
       ELSE

           "Z256_Manager".tOutputData.dMissionCode := "Z256_Manager".tInputData.dMissionCode;
           "Z256_Manager".tOutputData.rgxFireHeadON_OFF := "Z256_Manager".tInputData.rgxFireRequest;
           FOR #TMP_dIndex2 := 0 TO "CONST_dNumberOfHeadsCycle" DO
               "Z256_Manager".tOutputData.rgxDataToProcessInter[#TMP_dIndex2] := true;
           END_FOR;
           "Z256_Manager".tOutputData.dTargetLineValue_cmm := "Z256_Manager".tInputData.dMissionStart_cmm;

           #TMP_iReturn := "GP_BlockMoveStruct"(IN_iCount := DINT_TO_INT("CONST_dNumberOfHeads"),
                                                IN_iDestIndex := 0,
                                                IN_iSourceIndex := 0,
                                                INO_vDestArrayStruct := "Z256_Manager".tOutputData.rgdHeadsPositions_cmm,
                                                INO_vSourceArrayStruct := "Z256_Manager".tInputData.rgdHeadsPosition_cmm);
       END_IF;

       //Copy the values for the end       
       "Z256_Manager".rgtInterruptMissionTank[#TMP_dIndex].dMissionCode := "Z256_Manager".tInputData.dMissionCode;
       "Z256_Manager".rgtInterruptMissionTank[#TMP_dIndex].dMissionValue_cmm := "Z256_Manager".tInputData.dMissionEnd_cmm;
       FOR #TMP_dIndex3 := 0 TO "CONST_dNumberOfHeadsCycle" DO
           "Z256_Manager".rgtInterruptMissionTank[#TMP_dIndex].rgxFireRequest [#TMP_dIndex3] := 0;
       END_FOR;

       #TMP_iReturn := "GP_BlockMoveStruct"(IN_iCount := DINT_TO_INT("CONST_dNumberOfHeads"),
                                            IN_iDestIndex := 0,
                                            IN_iSourceIndex := 0,
                                            INO_vDestArrayStruct := "Z256_Manager".rgtInterruptMissionTank[#TMP_dIndex].rgdHeadsPositions_cmm,
                                            INO_vSourceArrayStruct := "Z256_Manager".tInputData.rgdHeadsPosition_cmm);

       //Increment the tank position
       "Z256_Manager".dInterruptNumMissionTank := #TMP_dIndex + 1;

       //------- END INSERT MISSION FOR INTERRUPT -----------

       //------- INSERT MISSION FOR OIL AND ARM -------------
       //Insert only the request head
       FOR #TMP_dIndex := 0 TO "CONST_dNumberOfHeadsCycle" DO

           //Insert on buffer only the fire on head
           IF "Z256_Manager".tInputData.rgxFireRequest[#TMP_dIndex] THEN

               //----------- OIL -------------------

               #TMP_dInsideIndex := "Z256_Manager".rgtOilList[#TMP_dIndex].dNumberOfElement;

               #TMP_xOutputMergeMission := 0;

               IF ("Z256_Manager".rgtOilList[#TMP_dIndex].dNumberOfElement > 0) THEN

                   #TMP_dDummy := "Z256_Manager".tInputData.dMissionStart_cmm - "Z256_Manager".rgtOilList[#TMP_dIndex].rgdRequestPosition_cmm[#TMP_dInsideIndex - 1];

                   IF ABS(#TMP_dDummy) <= "CONST_dFire_OnOff_MaxValue" THEN
                       //The difference is less than the maximum offset. Merge the mission
                       #TMP_dInsideIndex := #TMP_dInsideIndex - 1;
                   END_IF;

               ELSE

                   #TMP_dDummy := "Z256_Manager".tInputData.dMissionStart_cmm - "Z256_Manager".tOutputData.rgdOilRequestTarget_cmm[#TMP_dIndex];

                   IF ABS(#TMP_dDummy) <= "CONST_dFire_OnOff_MaxValue" THEN
                       //The difference is less than the maximum offset. Merge the mission
                       #TMP_xOutputMergeMission := 1;
                   END_IF;

               END_IF;

               //Copy the start value
               IF NOT #TMP_xOutputMergeMission THEN

                   "Z256_Manager".rgtOilList[#TMP_dIndex].rgdRequestPosition_cmm[#TMP_dInsideIndex] := "Z256_Manager".tInputData.dMissionStart_cmm;
                   "Z256_Manager".rgtOilList[#TMP_dIndex].rgdFireRequest[#TMP_dInsideIndex] := 1;
                   "Z256_Manager".rgtOilList[#TMP_dIndex].rgdMissionID[#TMP_dInsideIndex] := "Z256_Manager".tInputData.dMissionCode;


                   #TMP_dInsideIndex := #TMP_dInsideIndex + 1;

               ELSE
                   "Z256_Manager".tOutputData.rgxOilRequest[#TMP_dIndex] := 1;
                   "Z256_Manager".tOutputData.rgdOilRequestTarget_cmm[#TMP_dIndex] := "Z256_Manager".tInputData.dMissionStart_cmm;

               END_IF;
               //Copy the end value
               "Z256_Manager".rgtOilList[#TMP_dIndex].rgdRequestPosition_cmm[#TMP_dInsideIndex] := "Z256_Manager".tInputData.dMissionEnd_cmm;
               "Z256_Manager".rgtOilList[#TMP_dIndex].rgdFireRequest[#TMP_dInsideIndex] := 0;
               "Z256_Manager".rgtOilList[#TMP_dIndex].rgdMissionID[#TMP_dInsideIndex] := "Z256_Manager".tInputData.dMissionCode;


               "Z256_Manager".rgtOilList[#TMP_dIndex].dNumberOfElement := #TMP_dInsideIndex + 1;

               //----------- ARM -------------------

               #TMP_dInsideIndex := "Z256_Manager".rgtArmList[#TMP_dIndex].dNumberOfElement;

               #TMP_xOutputMergeMission := 0;

               IF ("Z256_Manager".rgtArmList[#TMP_dIndex].dNumberOfElement > 0) THEN

                   #TMP_dDummy := "Z256_Manager".tInputData.dMissionStart_cmm - "Z256_Manager".rgtArmList[#TMP_dIndex].rgdRequestPosition_cmm[#TMP_dInsideIndex - 1];

                   IF ABS(#TMP_dDummy) <= "CONST_dFire_OnOff_MaxValue" THEN
                       //The difference is less than the maximum offset. Merge the mission
                       #TMP_dInsideIndex := #TMP_dInsideIndex - 1;
                   END_IF;

               ELSE

                   #TMP_dDummy := "Z256_Manager".tInputData.dMissionStart_cmm - "Z256_Manager".tOutputData.rgdArmRequestTarget_cmm[#TMP_dIndex];

                   IF ABS(#TMP_dDummy) <= "CONST_dFire_OnOff_MaxValue" THEN
                       //The difference is less than the maximum offset. Merge the mission
                       #TMP_xOutputMergeMission := 1;

                   END_IF;

               END_IF;

               //Copy the start value
               IF NOT #TMP_xOutputMergeMission THEN

                   "Z256_Manager".rgtArmList[#TMP_dIndex].rgdRequestPosition_cmm[#TMP_dInsideIndex] := "Z256_Manager".tInputData.dMissionStart_cmm;
                   "Z256_Manager".rgtArmList[#TMP_dIndex].rgdFireRequest[#TMP_dInsideIndex] := 1;
                   "Z256_Manager".rgtArmList[#TMP_dIndex].rgdMissionID[#TMP_dInsideIndex] := "Z256_Manager".tInputData.dMissionCode;

                   #TMP_dInsideIndex := #TMP_dInsideIndex + 1;
               ELSE

                   "Z256_Manager".tOutputData.rgxArmRequest[#TMP_dIndex] := 1;
                   "Z256_Manager".tOutputData.rgdArmRequestTarget_cmm[#TMP_dIndex] := "Z256_Manager".tInputData.dMissionStart_cmm;

               END_IF;

               //Copy the end value
               "Z256_Manager".rgtArmList[#TMP_dIndex].rgdRequestPosition_cmm[#TMP_dInsideIndex] := "Z256_Manager".tInputData.dMissionEnd_cmm;
               "Z256_Manager".rgtArmList[#TMP_dIndex].rgdFireRequest[#TMP_dInsideIndex] := 0;
               "Z256_Manager".rgtArmList[#TMP_dIndex].rgdMissionID[#TMP_dInsideIndex] := "Z256_Manager".tInputData.dMissionCode;

               "Z256_Manager".rgtArmList[#TMP_dIndex].dNumberOfElement := #TMP_dInsideIndex + 1;

           END_IF;
       END_FOR;

       //Reset the mission request flag
       "Z256_Manager".tInputData.xNewMission := 0;
       "CM_Manager".ST_xNewMissionCPU0 := 0;
   END_IF;



   FOR #TMP_dIndex := 0 TO "CONST_dNumberOfHeadsCycle" DO

       //OIL MANAGER

       REPEAT

           #TMP_xCheckNext := 0;

           IF ("Z256_Manager".rgtOilList[#TMP_dIndex].dNumberOfElement > 0) THEN

               //We have one element, check the request.
               IF ("Z256_Manager".rgtOilList[#TMP_dIndex].rgdFireRequest[0] = 1) THEN
                   #TMP_dDummy := "Z256_Manager".rgtOilList[#TMP_dIndex].rgdRequestPosition_cmm[0] -
                   ("Z256_Manager".tInputData.rgdFireONReaction_ms[#TMP_dIndex] * REAL_TO_DINT("Encoder".AUX_rActualSpeedValue_cmm_ms)) +
                   "Z256_Manager".tInputData.rgdFireONDelayStart_cmm[#TMP_dIndex] +
                   ("Z256_Manager".tInputData.rgdOilDelayStart_ms[#TMP_dIndex] * REAL_TO_DINT("Encoder".AUX_rActualSpeedValue_cmm_ms));

               ELSE
                   #TMP_dDummy := "Z256_Manager".rgtOilList[#TMP_dIndex].rgdRequestPosition_cmm[0] -
                   ("Z256_Manager".tInputData.rgdFireOFFReaction_ms[#TMP_dIndex] * REAL_TO_DINT("Encoder".AUX_rActualSpeedValue_cmm_ms)) +
                   "Z256_Manager".tInputData.rgdFireOFFDelayEnd_cmm[#TMP_dIndex] +
                   ("Z256_Manager".tInputData.rgdOilDelayEnd_ms[#TMP_dIndex] * REAL_TO_DINT("Encoder".AUX_rActualSpeedValue_cmm_ms));
               END_IF;

               //If we are over, execute the request and take out the element. 
               #TMP_dLineOverlap := "Encoder".AUX_dActualEncoderValue_cmm - #TMP_dDummy;

               IF (#TMP_dLineOverlap >= 0) THEN

                   //Move the request to output
                   IF "Z256_Manager".rgtOilList[#TMP_dIndex].rgdFireRequest[0] = 1 THEN
                       "Z256_Manager".tOutputData.rgxOilRequest[#TMP_dIndex] := 1;
                       "Z256_Manager".tOutputData.rgdOilRequestTarget_cmm[#TMP_dIndex] := "Z256_Manager".rgtOilList[#TMP_dIndex].rgdRequestPosition_cmm[0];
                       "Z256_Manager".tOutputData.rgdOilRequestIDMission[#TMP_dIndex] := "Z256_Manager".rgtOilList[#TMP_dIndex].rgdMissionID[0];

                   ELSE
                       "Z256_Manager".tOutputData.rgxOilRequest[#TMP_dIndex] := 0;
                       "Z256_Manager".tOutputData.rgdOilRequestTarget_cmm[#TMP_dIndex] := "Z256_Manager".rgtOilList[#TMP_dIndex].rgdRequestPosition_cmm[0];
                       "Z256_Manager".tOutputData.rgdOilRequestIDMission[#TMP_dIndex] := "Z256_Manager".rgtOilList[#TMP_dIndex].rgdMissionID[0];

                   END_IF;

                   //Decrement the number of element
                   "Z256_Manager".rgtOilList[#TMP_dIndex].dNumberOfElement := "Z256_Manager".rgtOilList[#TMP_dIndex].dNumberOfElement - 1;

                   IF ("Z256_Manager".rgtOilList[#TMP_dIndex].dNumberOfElement > 0) THEN

                       //Shift up the array data
                       #TMP_iReturn := "GP_BlockMoveStruct"(IN_iCount :=DINT_TO_INT("Z256_Manager".rgtOilList[#TMP_dIndex].dNumberOfElement),
                                                            IN_iDestIndex := 0,
                                                            IN_iSourceIndex := 1,
                                                            INO_vDestArrayStruct := "Z256_Manager".rgtOilList[#TMP_dIndex].rgdFireRequest,
                                                            INO_vSourceArrayStruct := "Z256_Manager".rgtOilList[#TMP_dIndex].rgdFireRequest);

                       #TMP_iReturn := "GP_BlockMoveStruct"(IN_iCount := DINT_TO_INT("Z256_Manager".rgtOilList[#TMP_dIndex].dNumberOfElement),
                                                            IN_iDestIndex := 0,
                                                            IN_iSourceIndex := 1,
                                                            INO_vDestArrayStruct := "Z256_Manager".rgtOilList[#TMP_dIndex].rgdRequestPosition_cmm,
                                                            INO_vSourceArrayStruct := "Z256_Manager".rgtOilList[#TMP_dIndex].rgdRequestPosition_cmm);

                       #TMP_iReturn := "GP_BlockMoveStruct"(IN_iCount := DINT_TO_INT("Z256_Manager".rgtOilList[#TMP_dIndex].dNumberOfElement),
                                                            IN_iDestIndex := 0,
                                                            IN_iSourceIndex := 1,
                                                            INO_vDestArrayStruct := "Z256_Manager".rgtOilList[#TMP_dIndex].rgdMissionID,
                                                            INO_vSourceArrayStruct := "Z256_Manager".rgtOilList[#TMP_dIndex].rgdMissionID);

                       //Ask the system to check the next value, to avoid overlap
                       #TMP_xCheckNext := 1;
                   END_IF;

                   #TMP_dDummy := "Z256_Manager".rgtOilList[#TMP_dIndex].dNumberOfElement;
                   "Z256_Manager".rgtOilList[#TMP_dIndex].rgdRequestPosition_cmm[#TMP_dDummy] := 0;
                   "Z256_Manager".rgtOilList[#TMP_dIndex].rgdFireRequest[#TMP_dDummy] := 0;
                   "Z256_Manager".rgtOilList[#TMP_dIndex].rgdMissionID[#TMP_dDummy] := 0;

               END_IF;

           END_IF;

       UNTIL NOT #TMP_xCheckNext
       END_REPEAT;

       //ARM MANAGER

       REPEAT

           #TMP_xCheckNext := 0;

           IF ("Z256_Manager".rgtArmList[#TMP_dIndex].dNumberOfElement > 0) THEN

               //We have one element, check the request.
               IF ("Z256_Manager".rgtArmList[#TMP_dIndex].rgdFireRequest[0] = 1) THEN
                   #TMP_dDummy := ("Z256_Manager".rgtArmList[#TMP_dIndex].rgdRequestPosition_cmm[0] -
                   ("Z256_Manager".tInputData.rgdFireONReaction_ms[#TMP_dIndex] * REAL_TO_DINT("Encoder".AUX_rActualSpeedValue_cmm_ms))) +
                   "Z256_Manager".tInputData.rgdFireONDelayStart_cmm[#TMP_dIndex] -
                   ("Z256_Manager".tInputData.rgdArmONReaction_ms[#TMP_dIndex] * REAL_TO_DINT("Encoder".AUX_rActualSpeedValue_cmm_ms));

               ELSE
                   #TMP_dDummy := ("Z256_Manager".rgtArmList[#TMP_dIndex].rgdRequestPosition_cmm[0] -
                   ("Z256_Manager".tInputData.rgdFireOFFReaction_ms[#TMP_dIndex] * REAL_TO_DINT("Encoder".AUX_rActualSpeedValue_cmm_ms))) +
                   "Z256_Manager".tInputData.rgdFireOFFDelayEnd_cmm[#TMP_dIndex] -
                   ("Z256_Manager".tInputData.rgdArmOFFReaction_ms[#TMP_dIndex] * REAL_TO_DINT("Encoder".AUX_rActualSpeedValue_cmm_ms));
               END_IF;

               //If we are over, execute the request and take out the element. 
               #TMP_dLineOverlap := "Encoder".AUX_dActualEncoderValue_cmm - #TMP_dDummy;

               IF (#TMP_dLineOverlap >= 0) THEN

                   //Move the request to output
                   IF "Z256_Manager".rgtArmList[#TMP_dIndex].rgdFireRequest[0] = 1 THEN
                       "Z256_Manager".tOutputData.rgxArmRequest[#TMP_dIndex] := 1;
                       "Z256_Manager".tOutputData.rgdArmRequestTarget_cmm[#TMP_dIndex] := "Z256_Manager".rgtArmList[#TMP_dIndex].rgdRequestPosition_cmm[0];
                       "Z256_Manager".tOutputData.rgdArmRequestIDMission[#TMP_dIndex] := "Z256_Manager".rgtArmList[#TMP_dIndex].rgdMissionID[0];
                   ELSE
                       "Z256_Manager".tOutputData.rgxArmRequest[#TMP_dIndex] := 0;
                       "Z256_Manager".tOutputData.rgdArmRequestTarget_cmm[#TMP_dIndex] := "Z256_Manager".rgtArmList[#TMP_dIndex].rgdRequestPosition_cmm[0];
                       "Z256_Manager".tOutputData.rgdArmRequestIDMission[#TMP_dIndex] := 0;
                   END_IF;

                   //Decrement the number of element
                   "Z256_Manager".rgtArmList[#TMP_dIndex].dNumberOfElement := "Z256_Manager".rgtArmList[#TMP_dIndex].dNumberOfElement - 1;

                   IF ("Z256_Manager".rgtArmList[#TMP_dIndex].dNumberOfElement > 0) THEN

                       //Shift up the array data
                       #TMP_iReturn := "GP_BlockMoveStruct"(IN_iCount := DINT_TO_INT("Z256_Manager".rgtArmList[#TMP_dIndex].dNumberOfElement),
                                                            IN_iDestIndex := 0,
                                                            IN_iSourceIndex := 1,
                                                            INO_vDestArrayStruct := "Z256_Manager".rgtArmList[#TMP_dIndex].rgdFireRequest,
                                                            INO_vSourceArrayStruct := "Z256_Manager".rgtArmList[#TMP_dIndex].rgdFireRequest);

                       #TMP_iReturn := "GP_BlockMoveStruct"(IN_iCount := DINT_TO_INT("Z256_Manager".rgtArmList[#TMP_dIndex].dNumberOfElement),
                                                            IN_iDestIndex := 0,
                                                            IN_iSourceIndex := 1,
                                                            INO_vDestArrayStruct := "Z256_Manager".rgtArmList[#TMP_dIndex].rgdRequestPosition_cmm,
                                                            INO_vSourceArrayStruct := "Z256_Manager".rgtArmList[#TMP_dIndex].rgdRequestPosition_cmm);

                       #TMP_iReturn := "GP_BlockMoveStruct"(IN_iCount := DINT_TO_INT("Z256_Manager".rgtArmList[#TMP_dIndex].dNumberOfElement),
                                                            IN_iDestIndex := 0,
                                                            IN_iSourceIndex := 1,
                                                            INO_vDestArrayStruct := "Z256_Manager".rgtArmList[#TMP_dIndex].rgdMissionID,
                                                            INO_vSourceArrayStruct := "Z256_Manager".rgtArmList[#TMP_dIndex].rgdMissionID);

                       //Ask the system to check the next value, to avoid overlap
                       #TMP_xCheckNext := 1;
                   END_IF;

                   //Clear the array data
                   #TMP_dDummy := "Z256_Manager".rgtArmList[#TMP_dIndex].dNumberOfElement;
                   "Z256_Manager".rgtArmList[#TMP_dIndex].rgdRequestPosition_cmm[#TMP_dDummy] := 0;
                   "Z256_Manager".rgtArmList[#TMP_dIndex].rgdFireRequest[#TMP_dDummy] := 0;
                   "Z256_Manager".rgtArmList[#TMP_dIndex].rgdMissionID[#TMP_dDummy] := 0;


               END_IF;

           END_IF;

       UNTIL NOT #TMP_xCheckNext
       END_REPEAT;


   END_FOR;

   //---- INTERRUPT MANAGER ----
   //This part will prepare the output data for the interrupt
   #TMP_xDummy := false;
   FOR #TMP_dIndex3 := 0 TO "CONST_dNumberOfHeadsCycle" DO
       IF "Z256_Manager".tOutputData.rgxDataToProcessInter[#TMP_dIndex3] = TRUE THEN
           #TMP_xDummy := true;
       END_IF;
   END_FOR;

   IF #TMP_xDummy=FALSE THEN

       //Interrupt has no data to manage. Check the next mission
       IF ("Z256_Manager".dInterruptNumMissionTank > 0) THEN

           //This part is to prevent the moving of the head if some arming and oil are still
           //in progress. To allow the mission change:

           #TMP_xProcNextAllowed := 1;

           #TMP_xIsDiffent := 0;

           FOR #TMP_dIndex := 0 TO "CONST_dNumberOfHeadsCycle" DO

               IF "Z256_Manager".tOutputData.rgdHeadsPositions_cmm[#TMP_dIndex] <> "Z256_Manager".rgtInterruptMissionTank[0].rgdHeadsPositions_cmm[#TMP_dIndex] THEN

                   #TMP_xIsDiffent := 1;
                   EXIT;

               END_IF;

           END_FOR;

           IF #TMP_xIsDiffent THEN
               FOR #TMP_dIndex := 0 TO "CONST_dNumberOfHeadsCycle" DO


                   IF "Z256_Manager".tOutputData.rgdArmRequestIDMission[#TMP_dIndex] <> 0 AND 
                       "Z256_Manager".tOutputData.rgdArmRequestIDMission[#TMP_dIndex] < "Z256_Manager".tOutputData.dMissionCode THEN;

                       //TMP_xProcNextAllowed := 0;
                   END_IF;



                   //           IF ("Z256_Manager".rgtArmList[#TMP_dIndex].dNumberOfElement > 0) AND ("Z256_Manager".rgtArmList[#TMP_dIndex].rgdMissionID[0] = "Z256_Manager".tOutputData.dMissionCode) AND
                   //               ("Z256_Manager".rgtArmList[#TMP_dIndex].rgdMissionID[0] <> "Z256_Manager".rgtInterruptMissionTank[0].dMissionCode) THEN

                   //              #TMP_xProcNextAllowed := 0;

                   //           END_IF;

                   //         IF ("Z256_Manager".rgtOilList[#TMP_dIndex].dNumberOfElement > 0) AND ("Z256_Manager".rgtOilList[#TMP_dIndex].rgdMissionID[0] = "Z256_Manager".tOutputData.dMissionCode) AND
                   //        ("Z256_Manager".rgtOilList[#TMP_dIndex].rgdMissionID[0] <> "Z256_Manager".rgtInterruptMissionTank[0].dMissionCode) THEN

                   //         #TMP_xProcNextAllowed := 0;

                   //       END_IF;


               END_FOR;
           END_IF;

           IF #TMP_xProcNextAllowed THEN

               //Take the first element and put in the output zone
               "Z256_Manager".tOutputData.xGateOpen := 0;

               "Z256_Manager".tOutputData.dMissionCode := "Z256_Manager".rgtInterruptMissionTank[0].dMissionCode;
               "Z256_Manager".tOutputData.rgxFireHeadON_OFF := "Z256_Manager".rgtInterruptMissionTank[0].rgxFireRequest;
               FOR #TMP_dIndex2 := 0 TO "CONST_dNumberOfHeadsCycle" DO
                   "Z256_Manager".tOutputData.rgxDataToProcessInter[#TMP_dIndex2] := true;
               END_FOR;
               "Z256_Manager".tOutputData.dTargetLineValue_cmm := "Z256_Manager".rgtInterruptMissionTank[0].dMissionValue_cmm;


               #TMP_iReturn := "GP_BlockMoveStruct"(IN_iCount := DINT_TO_INT("CONST_dNumberOfHeads"),
                                                    IN_iDestIndex := 0,
                                                    IN_iSourceIndex := 0,
                                                    INO_vDestArrayStruct := "Z256_Manager".tOutputData.rgdHeadsPositions_cmm,
                                                    INO_vSourceArrayStruct := "Z256_Manager".rgtInterruptMissionTank[0].rgdHeadsPositions_cmm);
               "Z256_Manager".tOutputData.rgdHeadsPositions_cmm[0]:= "Z256_Manager".rgtInterruptMissionTank[0].rgdHeadsPositions_cmm[0];


               //Mission copied, take out from buffer
               "Z256_Manager".dInterruptNumMissionTank := "Z256_Manager".dInterruptNumMissionTank - 1;

               IF ("Z256_Manager".dInterruptNumMissionTank > 0) THEN
                   #TMP_iReturn := "GP_BlockMoveStruct"(IN_iCount := DINT_TO_INT("Z256_Manager".dInterruptNumMissionTank),
                                                        IN_iDestIndex := 0,
                                                        IN_iSourceIndex := 1,
                                                        INO_vDestArrayStruct := "Z256_Manager".rgtInterruptMissionTank,
                                                        INO_vSourceArrayStruct := "Z256_Manager".rgtInterruptMissionTank);
               END_IF;

               //Clear the array data
               "Z256_Manager".rgtInterruptMissionTank["Z256_Manager".dInterruptNumMissionTank].dMissionCode := 0;
               "Z256_Manager".rgtInterruptMissionTank["Z256_Manager".dInterruptNumMissionTank].dMissionValue_cmm := 0;
               FOR #TMP_dIndex := 0 TO "CONST_dNumberOfHeadsCycle" DO
                   "Z256_Manager".rgtInterruptMissionTank["Z256_Manager".dInterruptNumMissionTank].rgxFireRequest [#TMP_dIndex] := 0;
               END_FOR;

               FOR #TMP_dIndex := 0 TO "CONST_dNumberOfHeadsCycle" DO
                   "Z256_Manager".rgtInterruptMissionTank["Z256_Manager".dInterruptNumMissionTank].rgdHeadsPositions_cmm[#TMP_dIndex] := 0;
               END_FOR;
           END_IF;
       END_IF;
   END_IF;

   #TMP_xDummy := false;
   FOR #TMP_dIndex2 := 0 TO "CONST_dNumberOfHeadsCycle" DO
       IF   "Z256_Manager".tOutputData.rgxDataToProcessInter[#TMP_dIndex2] = true THEN
           #TMP_xDummy := true;
       END_IF;
   END_FOR;
   //This part will calculate the fire ON threshold
   IF #TMP_xDummy AND (NOT "Z256_Manager".tOutputData.xGateOpen) THEN

       #TMP_xDummy := 0;

       FOR #TMP_dIndex := 0 TO "CONST_dNumberOfHeadsCycle" DO

           IF "Z256_Manager".tOutputData.rgxFireHeadON_OFF[#TMP_dIndex] THEN
               "Z256_Manager".tOutputData.rgdFireHeadThreshold_cmm[#TMP_dIndex] := ("Z256_Manager".tOutputData.dTargetLineValue_cmm + "Z256_Manager".tInputData.rgdFireONDelayStart_cmm[#TMP_dIndex]) -
               ("Z256_Manager".tInputData.rgdFireONReaction_ms[#TMP_dIndex] * REAL_TO_DINT("Encoder".AUX_rActualSpeedValue_cmm_ms));
           ELSE
               "Z256_Manager".tOutputData.rgdFireHeadThreshold_cmm[#TMP_dIndex] := ("Z256_Manager".tOutputData.dTargetLineValue_cmm + "Z256_Manager".tInputData.rgdFireOFFDelayEnd_cmm[#TMP_dIndex]) -
               ("Z256_Manager".tInputData.rgdFireOFFReaction_ms[#TMP_dIndex] * REAL_TO_DINT("Encoder".AUX_rActualSpeedValue_cmm_ms));
           END_IF;

           //Check if we are near the window. If we are (around 250mm before) i will open the interrupt

           #TMP_dDummy := "Encoder".AUX_dActualEncoderValue_cmm - "Z256_Manager".tOutputData.rgdFireHeadThreshold_cmm[#TMP_dIndex];

           IF (#TMP_dDummy >= -25000) THEN

               //The threshold is near the limits. Open the gate
               #TMP_xDummy := 1;
           END_IF;
       END_FOR;

       "Z256_Manager".tOutputData.xGateOpen := #TMP_xDummy;

   ELSE
       #TMP_xDummy := false;
       FOR #TMP_dIndex2 := 0 TO "CONST_dNumberOfHeadsCycle" DO
           IF "Z256_Manager".tOutputData.rgxDataToProcessInter[#TMP_dIndex2] = true THEN
               #TMP_xDummy := true;
           END_IF;
       END_FOR;
       IF ("Z256_Manager".tOutputData.xGateOpen) AND #TMP_xDummy=0 THEN

           //Reset the gate
           "Z256_Manager".tOutputData.xGateOpen := 0;

       END_IF;

   END_IF;


   //Reset cleaner
   //this part will reset all the information data, in order to give the system ready
   //for the next mission
   IF "Z256_Manager".tInputData.xSystemReset THEN

       "Z256_Manager".tInputData.xSystemReset := 0;

       //RESET OIL DATA
       #TMP_dSize := "GP_GetArraySize"("Z256_Manager".rgtOilList);
       FOR #TMP_dIndex := 0 TO #TMP_dSize - 1 DO

           "Z256_Manager".rgtOilList[#TMP_dIndex].dNumberOfElement := 0;

           #TMP_dSize2 := "GP_GetArraySize"("Z256_Manager".rgtOilList[#TMP_dIndex].rgdRequestPosition_cmm);

           FOR #TMP_dIndex2 := 0 TO #TMP_dSize2 - 1 DO
               "Z256_Manager".rgtOilList[#TMP_dIndex].rgdRequestPosition_cmm[#TMP_dIndex2] := 0;
           END_FOR;

           #TMP_dSize2 := "GP_GetArraySize"("Z256_Manager".rgtOilList[#TMP_dIndex].rgdFireRequest);

           FOR #TMP_dIndex2 := 0 TO #TMP_dSize2 - 1 DO
               "Z256_Manager".rgtOilList[#TMP_dIndex].rgdFireRequest[#TMP_dIndex2] := 0;
           END_FOR;

           #TMP_dSize2 := "GP_GetArraySize"("Z256_Manager".rgtOilList[#TMP_dIndex].rgdMissionID);

           FOR #TMP_dIndex2 := 0 TO #TMP_dSize2 - 1 DO
               "Z256_Manager".rgtOilList[#TMP_dIndex].rgdMissionID[#TMP_dIndex2] := 0;
           END_FOR;

       END_FOR;

       FOR #TMP_dIndex := 0 TO "CONST_dNumberOfHeadsCycle" DO
           "Z256_Manager".tOutputData.rgxOilRequest[#TMP_dIndex] := 0;
       END_FOR;

       //RESET ARM DATA
       #TMP_dSize := "GP_GetArraySize"("Z256_Manager".rgtArmList);
       FOR #TMP_dIndex := 0 TO #TMP_dSize - 1 DO

           "Z256_Manager".rgtArmList[#TMP_dIndex].dNumberOfElement := 0;

           #TMP_dSize2 := "GP_GetArraySize"("Z256_Manager".rgtArmList[#TMP_dIndex].rgdRequestPosition_cmm);

           FOR #TMP_dIndex2 := 0 TO #TMP_dSize2 - 1 DO
               "Z256_Manager".rgtArmList[#TMP_dIndex].rgdRequestPosition_cmm[#TMP_dIndex2] := 0;
           END_FOR;

           #TMP_dSize2 := "GP_GetArraySize"("Z256_Manager".rgtArmList[#TMP_dIndex].rgdFireRequest);

           FOR #TMP_dIndex2 := 0 TO #TMP_dSize2 - 1 DO
               "Z256_Manager".rgtArmList[#TMP_dIndex].rgdFireRequest[#TMP_dIndex2] := 0;
           END_FOR;

           #TMP_dSize := "GP_GetArraySize"("Z256_Manager".rgtArmList[#TMP_dIndex].rgdMissionID);

           FOR #TMP_dIndex2 := 0 TO #TMP_dSize2 - 1 DO
               "Z256_Manager".rgtArmList[#TMP_dIndex].rgdMissionID[#TMP_dIndex2] := 0;
           END_FOR;

       END_FOR;

       FOR #TMP_dIndex3 := 0 TO "CONST_dNumberOfHeadsCycle" DO
           "Z256_Manager".tOutputData.rgxArmRequest[#TMP_dIndex3] := 0;
       END_FOR;


       //RESET FIRE DATA
       #TMP_dSize := "GP_GetArraySize"("Z256_Manager".rgtInterruptMissionTank);

       "Z256_Manager".dInterruptNumMissionTank := 0;

       FOR #TMP_dIndex := 0 TO #TMP_dSize - 1 DO

           "Z256_Manager".rgtInterruptMissionTank[#TMP_dIndex].dMissionCode := 0;
           FOR #TMP_dIndex3 := 0 TO "CONST_dNumberOfHeadsCycle" DO
               "Z256_Manager".rgtInterruptMissionTank[#TMP_dIndex].rgxFireRequest[#TMP_dIndex3] := 0;
           END_FOR;
           "Z256_Manager".rgtInterruptMissionTank[#TMP_dIndex].dMissionValue_cmm := 0;

           #TMP_dSize2 := "GP_GetArraySize"("Z256_Manager".rgtInterruptMissionTank[#TMP_dIndex].rgdHeadsPositions_cmm);

           FOR #TMP_dIndex2 := 0 TO #TMP_dSize2 - 1 DO
               "Z256_Manager".rgtInterruptMissionTank[#TMP_dIndex].rgdHeadsPositions_cmm[#TMP_dIndex2] := 0;
           END_FOR;
       END_FOR;

       "Z256_Manager".tOutputData.dMissionCode := 0;
       FOR #TMP_dIndex3 := 0 TO "CONST_dNumberOfHeadsCycle" DO
           "Z256_Manager".tOutputData.rgxFireHeadON_OFF[#TMP_dIndex3] := 0;
       END_FOR;

       #TMP_xDummy := false;
       FOR #TMP_dIndex3 := 0 TO "CONST_dNumberOfHeadsCycle" DO
           "Z256_Manager".tOutputData.rgxDataToProcessInter[#TMP_dIndex3] := false;
       END_FOR;

       "Z256_Manager".tOutputData.xGateOpen := 0;
       "Z256_Manager".tOutputData.dTargetLineValue_cmm := 0;

       #TMP_dSize := "GP_GetArraySize"("Z256_Manager".tOutputData.rgdHeadsPositions_cmm);

       FOR #TMP_dIndex := 0 TO #TMP_dSize - 1 DO
           "Z256_Manager".tOutputData.rgdHeadsPositions_cmm[#TMP_dIndex] := 0;
       END_FOR;

       #TMP_dSize := "GP_GetArraySize"("Z256_Manager".tOutputData.rgdFireHeadThreshold_cmm);

       FOR #TMP_dIndex := 0 TO #TMP_dSize - 1 DO
           "Z256_Manager".tOutputData.rgdFireHeadThreshold_cmm[#TMP_dIndex] := 0;
       END_FOR;

       #TMP_dSize := "GP_GetArraySize"("Z256_Manager".tOutputData.rgdArmRequestTarget_cmm);


       #TMP_dSize := "GP_GetArraySize"("Z256_Manager".tOutputData.rgdArmRequestTarget_cmm);

       FOR #TMP_dIndex := 0 TO #TMP_dSize - 1 DO
           "Z256_Manager".tOutputData.rgdArmRequestTarget_cmm[#TMP_dIndex] := 0;
       END_FOR;

       #TMP_dSize := "GP_GetArraySize"("Z256_Manager".tOutputData.rgdOilRequestTarget_cmm);

       FOR #TMP_dIndex := 0 TO #TMP_dSize - 1 DO
           "Z256_Manager".tOutputData.rgdOilRequestTarget_cmm[#TMP_dIndex] := 0;
       END_FOR;

       #TMP_dSize := "GP_GetArraySize"("Z256_Manager".tOutputData.rgdArmRequestIDMission);

       FOR #TMP_dIndex := 0 TO #TMP_dSize - 1 DO
           "Z256_Manager".tOutputData.rgdArmRequestIDMission[#TMP_dIndex] := 0;
       END_FOR;

       #TMP_dSize := "GP_GetArraySize"("Z256_Manager".tOutputData.rgdOilRequestIDMission);

       FOR #TMP_dIndex := 0 TO #TMP_dSize - 1 DO
           "Z256_Manager".tOutputData.rgdOilRequestIDMission[#TMP_dIndex] := 0;
       END_FOR;


   END_IF;
END_FUNCTION

FUNCTION "M256M_SbrCalibratePosition" : Void   // FC6, SCL
{ S7_Optimized_Access := 'TRUE' }
VERSION : 0.1
   VAR_IN_OUT
      io_ST_xHeadReferredSwitch : Array[0.."CONST_dNumberOfHeadsCycle"] of Bool;
   END_VAR
   VAR_TEMP
      TMP_dIndex2 : DInt;
      TMP_dIndex : DInt;
      TMP_dGap_cmm : DInt;
   END_VAR
BEGIN
   ////--------------------------------------------------------------------------------------------------------------------
   //   Copyright (c)  Bottero Spa
   //--------------------------------------------------------------
   //   Routine: CalibratePosition                 
   //       Author: Alberto Cigliutti
   //   Created: <Date>
   //--------------------------------------------------------------
   //   Description: This function will calibrate the head position                
   //
   //   History:
   //
   ////--------------------------------------------------------------------------------------------------------------------

   FOR #TMP_dIndex := 0 TO "Z256_hmi".tHMW.dNumberOfLites - 1 DO

       //This operatio will do in this way.
       //The head of the first cut will be used as a reference.
       //The best way is to use the head #1 to to this job.
       //If the position is not correct, the function will change the home position of the head and all the heads
       //next the corrected one. This in order to give the same position.

       #TMP_dGap_cmm := "Z256_hmi".tHMW.rgdCutWidthReal_cmm[#TMP_dIndex] - "Z256_hmi".tHMW.rgdCutWidthTeo_cmm[#TMP_dIndex];

       //Positive value, mean that the real width is bigger than the request. That means we need to put the home position more near the center
       // in case of head with home on operator side. In case of head with home on opposite we need to put the home more far then the center

       FOR #TMP_dIndex2 := "Z256_hmi".tHMW.rgdHeadSelected[#TMP_dIndex + 1] - 1 TO "CONST_dNumberOfHeadsCycle" DO

           "M256_Manag_IDB".M256M_IDB[#TMP_dIndex2].tHMR.dHeadHomePositions_cmm := "M256_Manag_IDB".M256M_IDB[#TMP_dIndex2].tHMR.dHeadHomePositions_cmm + #TMP_dGap_cmm;

       END_FOR;

       //Operation done. Put the same value as request
       "Z256_hmi".tHMW.rgdCutWidthReal_cmm[#TMP_dIndex] := "Z256_hmi".tHMW.rgdCutWidthTeo_cmm[#TMP_dIndex];

   END_FOR;

   //Force the heads homing
   FOR #TMP_dIndex := 0 TO "CONST_dNumberOfHeadsCycle" DO
       #io_ST_xHeadReferredSwitch[#TMP_dIndex] := 0;
   END_FOR;
END_FUNCTION

FUNCTION "INPUT" : Void   // FC7, LAD
{ S7_Optimized_Access := 'TRUE' }
VERSION : 0.1
   VAR_TEMP
      iRetVal0 : Int;
      iRetVal1 : Int;
      wRetVal : Word;
   END_VAR
BEGIN

REGION Network 1 (SCL): Counter card
   "i.1B160AP1.CounterCardStatus" := "i.1B160AP1.CounterCardStatus":P;
   "i.1B160AP1.CounterActualValue" := "i.1B160AP1.CounterActualValue":P;
   "i.1B160AP1.CaptureValue" := "i.1B160AP1.CaptureValue":P;
   "i.1B160AP1.FrequencyActualValue" := "i.1B160AP1.FrequencyActualValue":P;

   "Encoder".INPUT_dEncoderCounter_count := DWORD_TO_DINT("i.1B160AP1.CounterActualValue");
   "Encoder".INPUT_dMeterPulseValue_count := DWORD_TO_DINT("i.1B160AP1.CaptureValue");
   "Encoder".INPUT_dFrequencyCounter_Hz := REAL_TO_DINT("i.1B160AP1.FrequencyActualValue");
   "Encoder".INPUT_xMeterPulseArrived := "i.1B160AP1.Event_Capture";
   "Encoder".INPUT_xResetEventAcknowledge := "i.1B160AP1.Res_Event_Ack";
END_REGION

REGION Network 2 (SCL): MCC1256
   "Z256".INPUT_xInputCtrlCabinetON := "i.1B160AP1.1B18-2L+.PowerSupplyInputControlCabinetON";
   "Z256".INPUT_xInputPowerSupplyON := "i.1B160AP1.1B18-3L+.InputInstallationPowerSupplyON";
   "Z256".INPUT_xAnomalyPower120_240 := "i.1B160AP1.1B11QF1/2.AnomalyPowerSupplies230V";
   "Z256".INPUT_xPowerSupply24vLogic1 := "i.1B160AP1.1B18QF2.PowerSupply24VLogic";
   "Z256".INPUT_xPowerSupply24vLogic2 := "i.1B160AP1.1B18QF3.PowerSupply24VLogic";
   "Z256".INPUT_xPowerSupply24vLogic3 := "i.1B160AP1.1B20QF2.PowerSupply24VLogic";
   "Z256".INPUT_xPowerSupply24vLogic4 := "i.1B160AP1.1B20QF3.PowerSupply24VLogic";
   "Z256".INPUT_xPowerSupply24vLogic5 := TRUE;

   "Z256".INPUT_xMainEmergencyON := "i.1B160AP1.1B122KE1.MainEmergencyON";
   "Z256".INPUT_xLocalEmergencyON := TRUE;
   "Z256".INPUT_xProtSupply36v_1 := "i.1B160AP1.1B41QF1.ProtectionPowerSupply36V_Motor_1-4";
   "Z256".INPUT_xProtMotorLC_1 := "i.1B160AP1.1B41QF2.ProtectionPowerSupplyMotorsYcut_1-4";
   "Z256".INPUT_xProtSupply36v_2 := "i.1B160AP1.1B42QF1.ProtectionPowerSupply36V_Motor_5-8";
   "Z256".INPUT_xProtMotorLC_2 := "i.1B160AP1.1B42QF2.ProtectionPowerSupplyMotorsYcut_5-8";

   "M256_Manag_IDB".M256M_IDB[0].INPUT_xCarriageOverload := "i.1B160AP1.1B51QM1.ProtectionCarriageTranslation";
   "M256_Manag_IDB".M256M_IDB[1].INPUT_xCarriageOverload := "i.1B160AP1.1B52QM1.ProtectionCarriageTranslation";
   "M256_Manag_IDB".M256M_IDB[2].INPUT_xCarriageOverload := "i.1B160AP1.1B53QM1.ProtectionCarriageTranslation";
   "M256_Manag_IDB".M256M_IDB[3].INPUT_xCarriageOverload := "i.1B160AP1.1B54QM1.ProtectionCarriageTranslation";
   "M256_Manag_IDB".M256M_IDB[4].INPUT_xCarriageOverload := "i.1B160AP1.1B55QM1.ProtectionCarriageTranslation";
   "M256_Manag_IDB".M256M_IDB[5].INPUT_xCarriageOverload := "i.1B160AP1.1B56QM1.ProtectionCarriageTranslation";
   "M256_Manag_IDB".M256M_IDB[6].INPUT_xCarriageOverload := "i.1B160AP1.1B57QM1.ProtectionCarriageTranslation";
   "M256_Manag_IDB".M256M_IDB[7].INPUT_xCarriageOverload := "i.1B160AP1.1B58QM1.ProtectionCarriageTranslation";

   "Z256".INPUT_xOperatorOverstroke := "M256_Manag_IDB".M256M_IDB[0].Axis_Ref.x_IO_4;
   "Z256".INPUT_xOppoOperatorOverstroke := "M256_Manag_IDB".M256M_IDB[4].Axis_Ref.x_IO_4;
END_REGION

REGION Network 3 (SCL): 300A1 / 400A1
   "Z256".INPUT_xLocalEmergency_Cabinet := 0;
   "Z256".INPUT_xLocalEmergency_SB1 :="i.1B160AP1.M217B1SB1.LocalEmergency";
   "Z256".INPUT_xLocalEmergency_SB2 :="i.1B160AP1.M217B1SB2.LocalEmergency";
   "Z256".INPUT_xResetLocalEmergency :=  FALSE;

   "M256_Manag_IDB".M256A_IDB[0].INPUT_xHeadsUpIstan := "i.1B160AP1.M217B1SB3_SB4.HeadsUpIstantaneous" ;
   "M256_Manag_IDB".M256A_IDB[1].INPUT_xHeadsUpIstan := "i.1B160AP1.M217B1SB3_SB4.HeadsUpIstantaneous" ;
   "M256_Manag_IDB".M256A_IDB[2].INPUT_xHeadsUpIstan := "i.1B160AP1.M217B1SB3_SB4.HeadsUpIstantaneous" ;
   "M256_Manag_IDB".M256A_IDB[3].INPUT_xHeadsUpIstan := "i.1B160AP1.M217B1SB3_SB4.HeadsUpIstantaneous" ;
   "M256_Manag_IDB".M256A_IDB[4].INPUT_xHeadsUpIstan := "i.1B160AP1.M217B1SB3_SB4.HeadsUpIstantaneous" ;
   "M256_Manag_IDB".M256A_IDB[5].INPUT_xHeadsUpIstan := "i.1B160AP1.M217B1SB3_SB4.HeadsUpIstantaneous" ;
   "M256_Manag_IDB".M256A_IDB[6].INPUT_xHeadsUpIstan := "i.1B160AP1.M217B1SB3_SB4.HeadsUpIstantaneous" ;
   "M256_Manag_IDB".M256A_IDB[7].INPUT_xHeadsUpIstan := "i.1B160AP1.M217B1SB3_SB4.HeadsUpIstantaneous" ;
END_REGION

REGION Network 4 (SCL): Head #1
   "M256_Manag_IDB".M256F_IDB[0].INPUT_xPressureDec := "i.1B411AP1.1B411SA1.Head1.CuttingPressure-";
   "M256_Manag_IDB".M256A_IDB[0].INPUT_xCarriageInWorkPosition := "i.1B411AP1.1B411SQ1.Head1.CarriageHeadWorkPosition";
   "M256_Manag_IDB".M256F_IDB[0].INPUT_xPressureInc := "i.1B411AP1.1B411SA1.Head1.CuttingPressure+";
   "Z256".INPUT_rgxHeadsInProduction[0] := "i.1B411AP1.1B411SA2.Head1.ProductionON";
   "M256_Manag_IDB".M256F_IDB[0].INPUT_xForceFiring := 0;
   "M256_Manag_IDB".M256A_IDB[0].INPUT_xForceArming := 0;
   "M256_Manag_IDB".M256M_IDB[0].INPUT_xBrakeRelease := FALSE;
   "M256_Manag_IDB".M256M_IDB[0].INPUT_xOverstroke := TRUE;//"i.1B410AP1.1B291KA1.Head1-2.CarriageTraslationAntiCollision";
END_REGION

REGION Network 5 (SCL): Head #2
   "M256_Manag_IDB".M256F_IDB[1].INPUT_xPressureDec := "i.1B412AP1.1B412SA1.Head2.CuttingPressure-";
   "M256_Manag_IDB".M256A_IDB[1].INPUT_xCarriageInWorkPosition := "i.1B412AP1.1B412SQ1.Head2.CarriageHeadWorkPosition";
   "M256_Manag_IDB".M256F_IDB[1].INPUT_xPressureInc := "i.1B412AP1.1B412SA1.Head2.CuttingPressure+";
   "Z256".INPUT_rgxHeadsInProduction[1] := "i.1B412AP1.1B412SA2.Head2.ProductionON";
   "M256_Manag_IDB".M256F_IDB[1].INPUT_xForceFiring := 0;
   "M256_Manag_IDB".M256A_IDB[1].INPUT_xForceArming := 0;
   "M256_Manag_IDB".M256M_IDB[1].INPUT_xBrakeRelease := FALSE;
   "M256_Manag_IDB".M256M_IDB[1].INPUT_xOverstroke := TRUE;//"i.1B410AP1.1B291KA2.Head2-3.CarriageTraslationAntiCollision";
END_REGION

REGION Network 6 (SCL): Head #3
   "M256_Manag_IDB".M256F_IDB[2].INPUT_xPressureDec := "i.1B413AP1.1B413SA1.Head3.CuttingPressure-";
   "M256_Manag_IDB".M256A_IDB[2].INPUT_xCarriageInWorkPosition := "i.1B413AP1.1B413SQ1.Head3.CarriageHeadWorkPosition";
   "M256_Manag_IDB".M256F_IDB[2].INPUT_xPressureInc := "i.1B413AP1.1B413SA1.Head3.CuttingPressure+";
   "Z256".INPUT_rgxHeadsInProduction[2] := "i.1B413AP1.1B413SA2.Head3.ProductionON";
   "M256_Manag_IDB".M256F_IDB[2].INPUT_xForceFiring := 0;
   "M256_Manag_IDB".M256A_IDB[2].INPUT_xForceArming := 0;
   "M256_Manag_IDB".M256M_IDB[2].INPUT_xBrakeRelease := FALSE;
   "M256_Manag_IDB".M256M_IDB[2].INPUT_xOverstroke := TRUE;//"i.1B410AP1.1B291KA3.Head3-4.CarriageTraslationAntiCollision";
END_REGION

REGION Network 7 (SCL): Head #4
   "M256_Manag_IDB".M256F_IDB[3].INPUT_xPressureDec :="i.1B414AP1.1B414SA1.Head4.CuttingPressure-";
   "M256_Manag_IDB".M256A_IDB[3].INPUT_xCarriageInWorkPosition := "i.1B414AP1.1B414SQ1.Head4.CarriageHeadWorkPosition";
   "M256_Manag_IDB".M256F_IDB[3].INPUT_xPressureInc := "i.1B414AP1.1B414SA1.Head4.CuttingPressure+";
   "Z256".INPUT_rgxHeadsInProduction[3] := "i.1B414AP1.1B414SA2.Head4.ProductionON";
   "M256_Manag_IDB".M256F_IDB[3].INPUT_xForceFiring := 0;
   "M256_Manag_IDB".M256A_IDB[3].INPUT_xForceArming := 0;
   "M256_Manag_IDB".M256M_IDB[3].INPUT_xBrakeRelease := FALSE;
   "M256_Manag_IDB".M256M_IDB[3].INPUT_xOverstroke := TRUE;//"i.1B410AP1.1B291KA4.Head4-5.CarriageTraslationAntiCollision";
END_REGION

REGION Network 8 (SCL): Head #5
   "M256_Manag_IDB".M256F_IDB[4].INPUT_xPressureDec := "i.1B415AP1.1B415SA1.Head5.CuttingPressure-";
   "M256_Manag_IDB".M256A_IDB[4].INPUT_xCarriageInWorkPosition := "i.1B415AP1.1B415SQ1.Head5.CarriageHeadWorkPosition";
   "M256_Manag_IDB".M256F_IDB[4].INPUT_xPressureInc := "i.1B415AP1.1B415SA1.Head5.CuttingPressure+";
   "Z256".INPUT_rgxHeadsInProduction[4] :="i.1B415AP1.1B415SA2.Head5.ProductionON";
   "M256_Manag_IDB".M256F_IDB[4].INPUT_xForceFiring := 0;
   "M256_Manag_IDB".M256A_IDB[4].INPUT_xForceArming := 0;
   "M256_Manag_IDB".M256M_IDB[4].INPUT_xBrakeRelease := FALSE;
   "M256_Manag_IDB".M256M_IDB[4].INPUT_xOverstroke := TRUE;//"i.1B410AP1.1B291KA5.Head5-6.CarriageTraslationAntiCollision";
END_REGION

REGION Network 9 (SCL): Head #6 / Head #5
   "M256_Manag_IDB".M256F_IDB[5].INPUT_xPressureDec := "i.1B416AP1.1B416SA1.Head6.CuttingPressure-";
   "M256_Manag_IDB".M256A_IDB[5].INPUT_xCarriageInWorkPosition := "i.1B416AP1.1B416SQ1.Head6.CarriageHeadWorkPosition";
   "M256_Manag_IDB".M256F_IDB[5].INPUT_xPressureInc := "i.1B416AP1.1B416SA1.Head6.CuttingPressure+";
   "Z256".INPUT_rgxHeadsInProduction[5] :="i.1B416AP1.1B416SA2.Head6.ProductionON";
   "M256_Manag_IDB".M256F_IDB[5].INPUT_xForceFiring := 0;
   "M256_Manag_IDB".M256A_IDB[5].INPUT_xForceArming := 0;
   "M256_Manag_IDB".M256M_IDB[5].INPUT_xBrakeRelease := FALSE;
   "M256_Manag_IDB".M256M_IDB[5].INPUT_xOverstroke := TRUE;//"i.1B410AP1.1B291KA8.Head6-7.CarriageTraslationAntiCollision";
END_REGION

REGION Network 10 (SCL): Head #7 / Head #5
   "M256_Manag_IDB".M256F_IDB[6].INPUT_xPressureDec := "i.1B417AP1.1B417SA1.Head7.CuttingPressure-";
   "M256_Manag_IDB".M256A_IDB[6].INPUT_xCarriageInWorkPosition := "i.1B417AP1.1B417SQ1.Head7.CarriageHeadWorkPosition";
   "M256_Manag_IDB".M256F_IDB[6].INPUT_xPressureInc := "i.1B417AP1.1B417SA1.Head7.CuttingPressure+";
   "Z256".INPUT_rgxHeadsInProduction[6] :="i.1B417AP1.1B417SA2.Head7.ProductionON";
   "M256_Manag_IDB".M256F_IDB[6].INPUT_xForceFiring := 0;
   "M256_Manag_IDB".M256A_IDB[6].INPUT_xForceArming := 0;
   "M256_Manag_IDB".M256M_IDB[6].INPUT_xBrakeRelease := FALSE;
   "M256_Manag_IDB".M256M_IDB[6].INPUT_xOverstroke := TRUE;//"i.1B410AP1.1B291KA7.Head7-8.CarriageTraslationAntiCollision";
END_REGION

REGION Network 11 (SCL): Head #8 / Head #5
   "M256_Manag_IDB".M256F_IDB[7].INPUT_xPressureDec := "i.1B418AP1.1B418SA1.Head8.CuttingPressure-";
   "M256_Manag_IDB".M256A_IDB[7].INPUT_xCarriageInWorkPosition := "i.1B418AP1.1B418SQ1.Head8.CarriageHeadWorkPosition";
   "M256_Manag_IDB".M256F_IDB[7].INPUT_xPressureInc := "i.1B418AP1.1B418SA1.Head8.CuttingPressure+";
   "Z256".INPUT_rgxHeadsInProduction[7] :="i.1B418AP1.1B418SA2.Head8.ProductionON";
   "M256_Manag_IDB".M256F_IDB[7].INPUT_xForceFiring := 0;
   "M256_Manag_IDB".M256A_IDB[7].INPUT_xForceArming := 0;
   "M256_Manag_IDB".M256M_IDB[7].INPUT_xBrakeRelease := FALSE;
   "M256_Manag_IDB".M256M_IDB[7].INPUT_xOverstroke := TRUE;//"i.1B410AP1.1B291KA8.Head8-9.CarriageTraslationAntiCollision";
END_REGION

REGION Network 12 (SCL): IDevice
   "CM_IDEV_FromMainLine" := "i.IDeviceCPU0";
END_REGION
END_FUNCTION

